HMI tags "Default tag table"
   "Clock_0.5Hz" : Bool = PLC "Clock_0.5Hz", 1 s
   "messageView" : Bool, internal
   "buttonView" : Bool, internal
   "RPA10B_datablock_PA10B_fatal_error_state_lock" : Int, 1 s
   "RPA10B_datablock_PA10B_error_state_lock" : Int, 1 s
   "RPA10B_datablock_PA10B_big_fail_state_lock" : Int, 1 s
   "RPA10B_datablock_PA10B_fail_state_lock" : Int, 1 s
   "RPA10B_datablock_RPA10B_station_work_cyclus_state" : UInt, 1 s
   "RPA10R_LCDSwitchAutomat_Manual" : Bool = PLC "RPA10B_LCD_switch_manual_automat", 1 s
   "RPA10B_datablock_RPA10B_station_start" : Bool, 1 s
   "show_input_page" : Int, internal
   "PLC_datablock_stations_configuration" : Byte, 1 s
   "RPA10B_datablock_RPA10B_instruction_list_index" : Byte, 1 s
   "RPA20B_open_drawer" : Bool = PLC "RPA20B_open_drawer", 1 s
   "RPA10B_LCD_switch_manual_automat" : Bool = PLC "RPA10B_LCD_switch_manual_automat", 1 s
   "RPA10B_datablock_RPA10B_scanned_data" : String[254], 1 s
   "RPA10B_light" : Bool = PLC "RPA10B_light", 1 s
   "RPA10B_LCD_beacon_green" : Bool = PLC "RPA10B_LCD_beacon_green", 1 s
   "RPA10B_LCD_beacon_orange" : Bool = PLC "RPA10B_LCD_beacon_orange", 1 s
   "RPA10B_LCD_beacon_red" : Bool = PLC "RPA10B_LCD_beacon_red", 1 s
   "RPA10B_LCD_beacon_siren" : Bool = PLC "RPA10B_LCD_beacon_siren", 1 s
   "RPA10B_LCD_button_start" : Bool = PLC "RPA10B_LCD_button_start", 1 s
   "RPA10B_LCD_LED_blue_confirm_button" : Bool = PLC "RPA10B_LCD_LED_blue_confirm_button", 1 s
   "RPA10B_LCD_LED_green_start_button" : Bool = PLC "RPA10B_LCD_LED_green_start_button", 1 s
   "RPA10B_code_position_1" : Bool = PLC "RPA10B_code_position_1", 1 s
   "RPA10B_code_position_2" : Bool = PLC "RPA10B_code_position_2", 1 s
   "RPA10B_home_position_horizontal_carriage_sensor" : Bool = PLC "RPA10B_home_position_horizontal_carriage_sensor", 1 s
   "RPA10B_end_position_horizontal_carriage_sensor" : Bool = PLC "RPA10B_end_position_horizontal_carriage_sensor", 1 s
   "RPA10B_home_position_idler_carriage_sensor" : Bool = PLC "RPA10B_home_position_idler_carriage_sensor", 1 s
   "RPA10B_end_position_idler_carriage_sensor" : Bool = PLC "RPA10B_end_position_idler_carriage_sensor", 1 s
   "RPA10B_idler_presence_sensor" : Bool = PLC "RPA10B_idler_presence_sensor", 1 s
   "show_output_page" : Int, internal
   "input_output" : Bool, internal
   "RPA10B_vacuum_sensor" : Bool = PLC "RPA10B_vacuum_sensor", 1 s
   "RPA10B_lock_sensor" : Bool = PLC "RPA10B_lock_sensor", 1 s
   "RPA10B_unlock_sensor" : Bool = PLC "RPA10B_unlock_sensor", 1 s
   "RPA10B_blend_1_vacuum_fix_sensor" : Bool = PLC "RPA10B_blend_1_vacuum_fix_sensor", 1 s
   "RPA10B_blend_2_vacuum_fix_sensor" : Bool = PLC "RPA10B_blend_2_vacuum_fix_sensor", 1 s
   "RPA10B_LCD_button_confirm" : Bool = PLC "RPA10B_LCD_button_confirm", 1 s
   "RPA10B_primerbox_pad_sensor_left" : Bool = PLC "RPA10B_primerbox_pad_sensor_left", 1 s
   "RPA10B_primerbox_pad_sensor_right" : Bool = PLC "RPA10B_primerbox_pad_sensor_right", 1 s
   "RPA10B_primerbox_felt_sensor" : Bool = PLC "RPA10B_primerbox_felt_sensor", 1 s
   "RPA10B_primerbox_felt_presence_sensor" : Bool = PLC "RPA10B_primerbox_felt_presence_sensor", 1 s
   "RPA10B_primerbox_button_PAD_IS_CHANGED" : Bool = PLC "RPA10B_primerbox_button_PAD_IS_CHANGED", 1 s
   "RPA10B_primerbox_bottle_2" : Bool = PLC "RPA10B_primerbox_bottle_2", 1 s
   "RPA10B_primerbox_bottle_1" : Bool = PLC "RPA10B_primerbox_bottle_1", 1 s
   "RPA10B_EJ_1_vacuum_sensor" : Bool = PLC "RPA10B_EJ_1_vacuum_sensor", 1 s
   "RPA10B_EJ_2_vacuum_sensor" : Bool = PLC "RPA10B_EJ_2_vacuum_sensor", 1 s
   "RPA10B_universal_button_1" : Bool = PLC "RPA10B_universal_button_1", 1 s
   "RPA10B_universal_button_2" : Bool = PLC "RPA10B_universal_button_2", 1 s
   "RPA20B_belt_position_sensor" : Bool = PLC "RPA20B_belt_position_sensor", 1 s
   "RPA20B_blend_presence_sensor_1" : Bool = PLC "RPA20B_blend_presence_sensor_1", 1 s
   "RPA20B_blend_presence_sensor_2" : Bool = PLC "RPA20B_blend_presence_sensor_2", 1 s
   "RPA20B_drawer_position_sensor" : Bool = PLC "RPA20B_drawer_position_sensor", 1 s
   "RPA20B_drawer_lock_sensor" : Bool = PLC "RPA20B_drawer_lock_sensor", 1 s
   "RPA20B_drawer_unlock_sensor" : Bool = PLC "RPA20B_drawer_unlock_sensor", 1 s
   "RPA20B_ES_feedback" : Bool = PLC "RPA20B_ES_feedback", 1 s
   "RPA20B_lock_door_feedback" : Bool = PLC "RPA20B_lock_door_feedback", 1 s
   "RPA20B_manual_UP" : Bool = PLC "RPA20B_manual_UP", 1 s
   "RPA20B_manual_DOWN" : Bool = PLC "RPA20B_manual_DOWN", 1 s
   "RPA20B_manual_move" : Bool = PLC "RPA20B_manual_move", 1 s
   "RPA20B_unlock_button" : Bool = PLC "RPA20B_unlock_button", 1 s
   "RPA20B_button_back_1" : Bool = PLC "RPA20B_button_back_1", 1 s
   "RPA20B_button_back_2" : Bool = PLC "RPA20B_button_back_2", 1 s
   "RPA10B_primerbox_beacon_green" : Bool = PLC "RPA10B_primerbox_beacon_green", 1 s
   "RPA10B_primerbox_beacon_orange" : Bool = PLC "RPA10B_primerbox_beacon_orange", 1 s
   "RPA10B_primerbox_beacon_red" : Bool = PLC "RPA10B_primerbox_beacon_red", 1 s
   "RPA10B_primerbox_beacon_siren" : Bool = PLC "RPA10B_primerbox_beacon_siren", 1 s
   "RPA10B_primerbox_LED_green_ready" : Bool = PLC "RPA10B_primerbox_LED_green_ready", 1 s
   "RPA10B_primerbox_LED_green_felt" : Bool = PLC "RPA10B_primerbox_LED_green_felt", 1 s
   "RPA10B_primerbox_LED_green_bottle_1" : Bool = PLC "RPA10B_primerbox_LED_green_bottle_1", 1 s
   "RPA10B_primerbox_LED_green_bottle_2" : Bool = PLC "RPA10B_primerbox_LED_green_bottle_2", 1 s
   "RPA10B_primerbox_LED_red_NOT_READY" : Bool = PLC "RPA10B_primerbox_LED_red_NOT_READY", 1 s
   "RPA10B_primerbox_LED_orange_change_pad" : Bool = PLC "RPA10B_primerbox_LED_orange_change_pad", 1 s
   "RPA10B_vavle_aretation_unlock" : Bool = PLC "RPA10B_vavle_aretation_unlock", 1 s
   "RPA10B_vavle_aretation_lock" : Bool = PLC "RPA10B_vavle_aretation_lock", 1 s
   "RPA10B_vavle_seal_idler_unlock" : Bool = PLC "RPA10B_vavle_seal_idler_unlock", 1 s
   "RPA10B_vavle_seal_idler_lock" : Bool = PLC "RPA10B_vavle_seal_idler_lock", 1 s
   "RPA10B_EJ_1_vacuum_control" : Bool = PLC "RPA10B_EJ_1_vacuum_control", 1 s
   "RPA10B_EJ_2_vacuum_control" : Bool = PLC "RPA10B_EJ_2_vacuum_control", 1 s
   "RPA10B_EJ_1_eject" : Bool = PLC "RPA10B_EJ_1_eject", 1 s
   "RPA10B_EJ_2_eject" : Bool = PLC "RPA10B_EJ_2_eject", 1 s
   "RPA10B_vacuum_cleaner_switch" : Bool = PLC "RPA10B_vacuum_cleaner_switch", 1 s
   "RPA20B_open_door_LED_green" : Bool = PLC "RPA20B_open_door_LED_green", 1 s
   "RPA20B_button_back_LED_1" : Bool = PLC "RPA20B_button_back_LED_1", 1 s
   "RPA20B_button_back_LED_2" : Bool = PLC "RPA20B_button_back_LED_2", 1 s
   "RPA20B_valve_open_drawer" : Bool = PLC "RPA20B_valve_open_drawer", 1 s
   "RPA20B_valve_close_drawer" : Bool = PLC "RPA20B_valve_close_drawer", 1 s
   "RPA20B_motor_down" : Bool = PLC "RPA20B_motor_down", 1 s
   "RPA20_motor_up" : Bool = PLC "RPA20_motor_up", 1 s
   "manual_page_switch" : Int, internal
   "RPA10B_datablock_RPA10B_show_pad_left" : Bool, 1 s
   "RPA10B_datablock_RPA10B_show_pad_right" : Bool, 1 s
   "RPA10B_datablock_RPA10_B_show_home" : Bool, 1 s
   "RPA10B_datablock_pa10B_bottle_cyclus_replace" : UInt, 1 s
   "RPA10B_datablock_pa10B_bottle_timing" : Time, 1 s

text list "PA10B_instructionList": 0 ''; 1 ''; 2 ''; 4 ''; 6 ''; 7 ''; 8 ''; 3 ''; 5 ''; 9 ''; 11 ''; 12 ''; 13 ''; 14 ''; 15 ''; 16 ''; 17 ''; 18 ''; 19 ''; 20 ''; 21 ''; 22 ''; 23 ''; 24 ''; 25 ''; 26 ''; 27 ''; 28 ''; 29 ''; 30 ''; 31 ''; 70 ''

text list "PA10B_fatal_error_list": 150 ''; 1100 ''

text list "pa10B_fail_list": 150 ''; 303 ''; 304 ''; 203 ''; 204 ''; 205 ''; 180 ''

text list "PA10B_error_list": 1000 ''; 400 ''; 401 ''; 402 ''; 403 ''

text list "PA10B_big_fail_list": 305 ''; 205 ''; 169 ''

text list "PA10B_station_variant_choose": 0 ''; 1 ''; 2 ''; 3 ''

screen "Home" 800x480
   TextField "Text field_3" at 325,5 size 300x40
   TextField "Text field_2" at 2,85 size 70x40
   TextField "Text field_5" at 335,130 size 130x25
   TextField "Text field_6" at 20,171 size 330x22
   TextField "Text field_7" at 20,201 size 330x22
   TextField "Text field_8" at 20,231 size 330x22
   TextField "Text field_9" at 20,261 size 330x22
   TextField "Text field_10" at 20,291 size 330x22
   TextField "Text field_11" at 20,321 size 330x22
   TextField "Text field_12" at 20,351 size 330x22
   TextField "Text field_13" at 20,381 size 330x22
   Button "Button_1" at 640,420 size 80x60
   Button "HmiScreenItemData_1" at 0,420 size 80x60
   Button "HmiScreenItemData_2" at 400,420 size 80x60
   Button "Button_2" at 560,420 size 80x60
   Button "Button_6" at 720,420 size 80x60
   DateTimeField "Date/time field_1" at 650,27 size 150x25
   DateTimeField "Date/time field_2" at 650,0 size 150x28
   TextField "Text field_1" at 0,0 size 300x50
   Button "HmiScreenItemData_3" at 240,420 size 80x60
   Button "HmiScreenItemData_4" at 320,420 size 80x60
   Button "Button_3" at 480,420 size 80x60
   Button "HmiScreenItemData_5" at 80,420 size 80x60
   Button "HmiScreenItemData_6" at 160,420 size 80x60
   IOField "I/O field_1" at 73,85 size 70x40
   Button "Button_11" at 0,420 size 80x60
   Button "Button_12" at 80,420 size 80x60
   Button "Button_13" at 160,420 size 80x60
   Button "Button_14" at 240,420 size 80x60
   Button "Button_15" at 320,420 size 80x60
   Button "Button_16" at 400,420 size 80x60
   Button "Button_17" at 480,420 size 80x60
   Button "Button_18" at 560,420 size 80x60
   Button "Button_19" at 640,420 size 80x60
   Button "Button_20" at 720,420 size 80x60
   TextField "Text field_22" at 64,67 size 129x22
   AlarmView "Alarm view_1" at 60,90 size 680x320
   Button "Button_9" at 715,65 size 25x25
   TextField "Text field_37" at 360,54 size 120x25

screen "I0-State" 800x480
   TextField "Text field_3" at 325,5 size 300x40
   Button "Button_1" at 640,420 size 80x60
   Button "Button_4" at 160,420 size 80x60
   Button "HmiScreenItemData_3" at 400,420 size 80x60
   Button "Button_2" at 560,420 size 80x60
   Button "Button_6" at 720,420 size 80x60
   Button "HmiScreenItemData_2" at 240,420 size 80x60
   Button "HmiScreenItemData_4" at 320,420 size 80x60
   TextField "Text field_1" at 0,0 size 300x50
   DateTimeField "Date/time field_2" at 650,0 size 150x28
   DateTimeField "Date/time field_1" at 650,27 size 150x25
   Button "HmiScreenItemData_1" at 0,420 size 80x60
   Button "Button_3" at 480,420 size 80x60
   Button "Button_5" at 80,420 size 80x60
   Button "input_back" at 20,52 size 90x25
   Button "input_next" at 690,52 size 90x25
   Button "output_back" at 20,52 size 90x25
   Button "output_next" at 690,52 size 90x25
   TextField "Text field_2" at 20,85 size 330x22
   TextField "Text field_4" at 20,114 size 330x22
   TextField "Text field_5" at 20,144 size 330x22
   TextField "Text field_6" at 20,174 size 330x22
   TextField "Text field_13" at 20,204 size 330x22
   TextField "Text field_14" at 20,232 size 330x22
   TextField "Text field_15" at 20,260 size 330x22
   TextField "Text field_16" at 20,288 size 330x22
   TextField "Text field_17" at 20,316 size 330x22
   TextField "Text field_18" at 20,344 size 330x22
   TextField "Text field_19" at 19,374 size 330x22
   TextField "Text field_20" at 387,86 size 330x22
   TextField "Text field_21" at 387,115 size 330x22
   TextField "Text field_22" at 387,144 size 330x22
   TextField "Text field_23" at 387,173 size 330x22
   TextField "Text field_24" at 387,202 size 330x22
   TextField "Text field_26" at 387,231 size 330x22
   TextField "Text field_27" at 387,260 size 330x22
   TextField "Text field_28" at 387,289 size 330x22
   TextField "Text field_29" at 387,318 size 330x22
   TextField "Text field_30" at 387,347 size 330x22
   TextField "Text field_31" at 387,376 size 330x22
   Button "Button_11" at 0,420 size 80x60
   Button "Button_12" at 80,420 size 80x60
   Button "Button_13" at 160,420 size 80x60
   Button "Button_14" at 240,420 size 80x60
   Button "Button_15" at 320,420 size 80x60
   Button "Button_16" at 400,420 size 80x60
   Button "Button_17" at 480,420 size 80x60
   Button "Button_18" at 560,420 size 80x60
   Button "Button_19" at 640,420 size 80x60
   Button "Button_20" at 720,420 size 80x60
   TextField "Text field_25" at 64,67 size 129x22
   AlarmView "Alarm view_1" at 60,90 size 680x320
   Button "Button_9" at 715,65 size 25x25
   TextField "Text field_7" at 20,85 size 330x22
   TextField "Text field_8" at 19,115 size 330x22
   TextField "Text field_9" at 19,145 size 330x22
   TextField "Text field_10" at 19,175 size 330x22
   TextField "Text field_11" at 20,205 size 330x22
   TextField "Text field_12" at 20,235 size 330x22
   TextField "Text field_50" at 20,263 size 330x22
   TextField "Text field_51" at 20,291 size 330x22
   TextField "Text field_52" at 20,319 size 330x22
   TextField "Text field_53" at 20,347 size 330x22
   TextField "Text field_54" at 20,375 size 330x22
   TextField "Text field_55" at 387,86 size 330x22
   TextField "Text field_56" at 386,116 size 330x22
   TextField "Text field_57" at 386,146 size 330x22
   TextField "Text field_58" at 386,176 size 330x22
   TextField "Text field_59" at 387,206 size 330x22
   TextField "Text field_60" at 387,236 size 330x22
   TextField "Text field_61" at 387,264 size 330x22
   TextField "Text field_62" at 387,292 size 330x22
   TextField "Text field_63" at 387,320 size 330x22
   TextField "Text field_64" at 387,348 size 330x22
   TextField "Text field_65" at 387,376 size 330x22
   TextField "Text field_32" at 20,85 size 330x22
   TextField "Text field_33" at 20,114 size 330x22
   TextField "Text field_34" at 20,144 size 330x22
   TextField "Text field_35" at 20,174 size 330x22
   TextField "Text field_36" at 20,204 size 330x22
   TextField "Text field_37" at 20,232 size 330x22
   TextField "Text field_38" at 20,260 size 330x22
   TextField "Text field_39" at 20,288 size 330x22
   TextField "Text field_40" at 20,316 size 330x22
   TextField "Text field_41" at 20,344 size 330x22
   TextField "Text field_42" at 19,374 size 330x22
   TextField "Text field_43" at 387,86 size 330x22
   TextField "Text field_44" at 387,115 size 330x22
   TextField "Text field_45" at 387,144 size 330x22
   TextField "Text field_46" at 387,173 size 330x22
   TextField "Text field_47" at 387,202 size 330x22
   TextField "Text field_48" at 387,231 size 330x22
   TextField "Text field_49" at 387,260 size 330x22
   TextField "Text field_66" at 20,85 size 330x22
   TextField "Text field_67" at 19,115 size 330x22
   TextField "Text field_68" at 19,145 size 330x22
   TextField "Text field_69" at 19,175 size 330x22
   TextField "Text field_70" at 20,205 size 330x22
   TextField "Text field_71" at 20,235 size 330x22
   TextField "Text field_72" at 20,263 size 330x22
   TextField "Text field_73" at 20,291 size 330x22
   TextField "Text field_74" at 20,319 size 330x22
   TextField "Text field_75" at 20,347 size 330x22
   TextField "Text field_76" at 20,375 size 330x22
   TextField "Text field_77" at 360,54 size 120x25

screen "Main_page" 800x480
   Button "HmiScreenItemData_1" at 80,420 size 80x60
   TextField "Text field_2" at 0,85 size 800x25
   TextField "Text field_3" at 325,5 size 300x40
   Button "Button_4" at 480,420 size 80x60
   Button "Button_5" at 640,420 size 80x60
   Button "Button_1" at 0,420 size 80x60
   Button "HmiScreenItemData_2" at 160,420 size 80x60
   Button "Button_2" at 400,420 size 80x60
   Button "Button_3" at 560,420 size 80x60
   Button "Button_6" at 720,420 size 80x60
   Button "HmiScreenItemData_3" at 240,420 size 80x60
   Button "HmiScreenItemData_4" at 320,420 size 80x60
   TextField "Text field_1" at 0,0 size 300x50
   DateTimeField "Date/time field_2" at 650,0 size 150x28
   DateTimeField "Date/time field_1" at 650,27 size 150x25
   SymbolicIOField "Symbolic I/O field_1" at 10,110 size 780x90
   Button "HmiScreenItemData_5" at 80,420 size 80x60
   GraphicView "Graphic view_1" at 320,228 size 180x180
   Button "Button_11" at 0,420 size 80x60
   Button "Button_12" at 80,420 size 80x60
   Button "Button_13" at 160,420 size 80x60
   Button "Button_14" at 240,420 size 80x60
   Button "Button_15" at 320,420 size 80x60
   Button "Button_16" at 400,420 size 80x60
   Button "Button_17" at 480,420 size 80x60
   Button "Button_18" at 560,420 size 80x60
   Button "Button_19" at 640,420 size 80x60
   Button "Button_20" at 720,420 size 80x60
   TextField "Text field_5" at 64,67 size 129x22
   AlarmView "Alarm view_1" at 60,90 size 680x320
   Button "Button_9" at 715,65 size 25x25
   SymbolicIOField "Symbolic I/O field_2" at 0,170 size 800x110
   SymbolicIOField "Symbolic I/O field_3" at 0,170 size 800x110
   SymbolicIOField "Symbolic I/O field_4" at 0,170 size 800x110
   SymbolicIOField "Symbolic I/O field_5" at 0,170 size 800x110
   TextField "Text field_37" at 360,54 size 120x25
   GraphicView "Graphic view_2" at 260,225 size 345x187
   GraphicView "Graphic view_3" at 195,225 size 345x187
   TextField "Text field_4" at 306,290 size 237x43

screen "Manual" 800x480
   Button "Button_4" at 21,85 size 50x50
   Button "Button_12" at 730,85 size 50x50
   Button "Button_1" at 640,420 size 80x60
   Button "HmiScreenItemData_1" at 0,420 size 80x60
   Button "Button_2" at 560,420 size 80x60
   Button "Button_6" at 720,420 size 80x60
   Button "Button_34" at 400,420 size 80x60
   Button "HmiScreenItemData_3" at 240,420 size 80x60
   Button "HmiScreenItemData_4" at 320,420 size 80x60
   TextField "Text field_1" at 0,0 size 300x50
   DateTimeField "Date/time field_2" at 650,0 size 150x28
   DateTimeField "Date/time field_1" at 650,27 size 150x25
   Button "Button_5" at 160,420 size 80x60
   Button "Button_3" at 480,420 size 80x60
   Button "Button_7" at 80,420 size 80x60
   Button "Button_8" at 730,85 size 50x50
   Button "Button_9" at 21,85 size 50x50
   Button "Button_23" at 0,420 size 80x60
   Button "Button_24" at 80,420 size 80x60
   Button "Button_25" at 160,420 size 80x60
   Button "Button_26" at 240,420 size 80x60
   Button "Button_27" at 320,420 size 80x60
   Button "Button_28" at 400,420 size 80x60
   Button "Button_29" at 480,420 size 80x60
   Button "Button_30" at 560,420 size 80x60
   Button "Button_31" at 640,420 size 80x60
   Button "Button_32" at 720,420 size 80x60
   TextField "Text field_8" at 64,67 size 129x22
   AlarmView "Alarm view_1" at 60,90 size 680x320
   Button "Button_33" at 715,65 size 25x25
   Switch "Switch_8" at 300,149 size 64x32
   Switch "Switch_9" at 300,185 size 64x32
   Switch "Switch_10" at 300,221 size 64x32
   Switch "Switch_11" at 300,257 size 64x32
   Switch "Switch_12" at 300,293 size 64x32
   Switch "Switch_13" at 301,328 size 64x32
   TextField "Text field_15" at 76,149 size 200x32
   TextField "Text field_16" at 76,181 size 200x32
   TextField "Text field_17" at 75,221 size 200x32
   TextField "Text field_18" at 37,289 size 239x32
   TextField "Text field_19" at 26,257 size 250x32
   TextField "Text field_20" at 29,328 size 247x32
   Switch "Switch_1" at 634,148 size 64x32
   TextField "Text field_2" at 410,148 size 200x32
   Switch "Switch_2" at 301,363 size 64x32
   TextField "Text field_4" at 29,363 size 247x32
   Switch "Switch_3" at 634,184 size 64x32
   TextField "Text field_5" at 379,184 size 231x32
   Switch "Switch_4" at 635,220 size 64x32
   TextField "Text field_6" at 394,220 size 217x32
   Switch "Switch_5" at 636,256 size 64x32
   TextField "Text field_7" at 377,256 size 235x32
   Switch "Switch_6" at 637,292 size 64x32
   TextField "Text field_9" at 377,292 size 236x32
   Switch "Switch_7" at 638,328 size 64x32
   TextField "Text field_10" at 376,328 size 238x32
   Switch "Switch_14" at 639,364 size 64x32
   TextField "Text field_11" at 322,364 size 293x32
   Switch "Switch_15" at 300,149 size 64x32
   Switch "Switch_16" at 300,185 size 64x32
   Switch "Switch_17" at 300,221 size 64x32
   Switch "Switch_18" at 300,257 size 64x32
   Switch "Switch_19" at 300,293 size 64x32
   Switch "Switch_20" at 301,328 size 64x32
   TextField "Text field_12" at 55,149 size 221x32
   TextField "Text field_13" at 8,181 size 268x32
   TextField "Text field_14" at 44,221 size 231x32
   TextField "Text field_21" at 37,289 size 239x32
   TextField "Text field_22" at 26,257 size 250x32
   TextField "Text field_23" at 29,328 size 247x32
   Switch "Switch_21" at 634,148 size 64x32
   TextField "Text field_24" at 388,148 size 222x32
   Switch "Switch_22" at 301,363 size 64x32
   TextField "Text field_25" at 29,363 size 247x32
   Switch "Switch_23" at 634,184 size 64x32
   TextField "Text field_26" at 379,184 size 231x32
   Switch "Switch_24" at 635,220 size 64x32
   TextField "Text field_27" at 394,220 size 217x32
   Switch "Switch_25" at 636,256 size 64x32
   TextField "Text field_28" at 377,256 size 235x32
   Switch "Switch_26" at 637,292 size 64x32
   TextField "Text field_29" at 377,292 size 236x32
   Switch "Switch_27" at 638,328 size 64x32
   TextField "Text field_30" at 376,328 size 238x32
   Switch "Switch_28" at 639,364 size 64x32
   TextField "Text field_31" at 382,364 size 233x32
   Switch "Switch_29" at 300,149 size 64x32
   Switch "Switch_30" at 300,185 size 64x32
   Switch "Switch_31" at 300,221 size 64x32
   Switch "Switch_32" at 300,257 size 64x32
   Switch "Switch_33" at 300,293 size 64x32
   TextField "Text field_32" at 55,149 size 221x32
   TextField "Text field_33" at 8,181 size 268x32
   TextField "Text field_34" at 22,221 size 253x32
   TextField "Text field_35" at 37,289 size 239x32
   TextField "Text field_36" at 26,257 size 250x32
   TextField "Text field_37" at 360,54 size 120x25

screen "Scanner" 800x480
   IOField "I/O field_1" at 10,118 size 780x32
   TextField "Text field_2" at 10,86 size 141x22
   Button "Button_1" at 640,420 size 80x60
   Button "HmiScreenItemData_3" at 400,420 size 80x60
   Button "Button_2" at 560,420 size 80x60
   Button "Button_6" at 720,420 size 80x60
   DateTimeField "Date/time field_2" at 650,0 size 150x28
   TextField "Text field_1" at 0,0 size 300x50
   DateTimeField "Date/time field_1" at 650,27 size 150x25
   Button "HmiScreenItemData_2" at 240,420 size 80x60
   Button "HmiScreenItemData_4" at 320,420 size 80x60
   Button "HmiScreenItemData_1" at 0,420 size 80x60
   Button "HmiScreenItemData_5" at 480,420 size 80x60
   Button "HmiScreenItemData_6" at 160,420 size 80x60
   Button "HmiScreenItemData_7" at 80,420 size 80x60
   Button "Button_3" at 10,170 size 96x32
   Button "Button_11" at 0,420 size 80x60
   Button "Button_12" at 80,420 size 80x60
   Button "Button_13" at 160,420 size 80x60
   Button "Button_14" at 240,420 size 80x60
   Button "Button_15" at 320,420 size 80x60
   Button "Button_16" at 400,420 size 80x60
   Button "Button_17" at 480,420 size 80x60
   Button "Button_18" at 560,420 size 80x60
   Button "Button_19" at 640,420 size 80x60
   Button "Button_20" at 720,420 size 80x60
   TextField "Text field_5" at 64,67 size 129x22
   Button "Button_9" at 715,65 size 25x25
   AlarmView "Alarm view_1" at 60,90 size 680x320
   TextField "Text field_37" at 360,54 size 120x25

screen "System" 800x480
   TextField "Text field_3" at 325,5 size 300x40
   TextField "Text field_2" at 300,85 size 200x27
   Button "Button_4" at 10,290 size 170x60
   Button "Button_5" at 10,355 size 170x60
   Button "Button_7" at 213,290 size 170x60
   Button "Button_8" at 416,290 size 170x60
   Button "Button_9" at 620,290 size 170x60
   Button "Button_11" at 213,355 size 170x60
   Button "Button_12" at 416,355 size 170x60
   Button "Button_13" at 620,355 size 170x60
   AlarmView "Alarm view_1" at 10,113 size 780x172
   Button "HmiScreenItemData_1" at 0,420 size 80x60
   Button "Button_3" at 160,420 size 80x60
   Button "Button_14" at 240,420 size 80x60
   Button "Button_15" at 320,420 size 80x60
   Button "Button_16" at 400,420 size 80x60
   Button "Button_17" at 480,420 size 80x60
   Button "Button_2" at 560,420 size 80x60
   Button "Button_1" at 640,420 size 80x60
   Button "Button_6" at 720,420 size 80x60
   TextField "Text field_1" at 0,0 size 300x50
   DateTimeField "Date/time field_2" at 650,0 size 150x28
   DateTimeField "Date/time field_1" at 650,27 size 150x25
   Button "Button_10" at 80,420 size 80x60
   TextField "Text field_37" at 360,54 size 120x25

screen "chemical_setup" 800x480
   Button "HmiScreenItemData_3" at 400,420 size 80x60
   Button "Button_2" at 560,420 size 80x60
   Button "Button_6" at 720,420 size 80x60
   DateTimeField "Date/time field_2" at 650,0 size 150x28
   TextField "Text field_1" at 0,0 size 300x50
   DateTimeField "Date/time field_1" at 650,27 size 150x25
   Button "HmiScreenItemData_2" at 240,420 size 80x60
   Button "HmiScreenItemData_4" at 320,420 size 80x60
   Button "HmiScreenItemData_1" at 0,420 size 80x60
   Button "HmiScreenItemData_5" at 480,420 size 80x60
   Button "HmiScreenItemData_6" at 160,420 size 80x60
   Button "HmiScreenItemData_7" at 80,420 size 80x60
   IOField "I/O field_1" at 87,130 size 341x44
   IOField "I/O field_2" at 87,237 size 338x44
   TextField "Text field_2" at 85,100 size 137x25
   TextField "Text field_3" at 87,206 size 111x25
   TextField "Text field_4" at 435,245 size 93x20
   Button "Button_1" at 640,420 size 80x60
   Button "Button_11" at 0,420 size 80x60
   Button "Button_12" at 80,420 size 80x60
   Button "Button_13" at 160,420 size 80x60
   Button "Button_14" at 240,420 size 80x60
   Button "Button_15" at 320,420 size 80x60
   Button "Button_16" at 400,420 size 80x60
   Button "Button_17" at 480,420 size 80x60
   Button "Button_18" at 560,420 size 80x60
   Button "Button_19" at 640,420 size 80x60
   Button "Button_20" at 720,420 size 80x60
   TextField "Text field_5" at 64,67 size 129x22
   Button "Button_9" at 715,65 size 25x25
   AlarmView "Alarm view_1" at 60,90 size 680x320
   TextField "Text field_37" at 360,54 size 120x25

screen "User_management" 800x480
   TextField "Text field_3" at 325,5 size 300x40
   Button "HmiScreenItemData_1" at 0,420 size 80x60
   Button "Button_3" at 160,420 size 80x60
   Button "Button_14" at 240,420 size 80x60
   Button "Button_15" at 320,420 size 80x60
   Button "Button_16" at 400,420 size 80x60
   Button "Button_17" at 480,420 size 80x60
   Button "Button_2" at 560,420 size 80x60
   Button "Button_1" at 640,420 size 80x60
   TextField "Text field_1" at 0,0 size 300x50
   DateTimeField "Date/time field_2" at 650,0 size 150x28
   DateTimeField "Date/time field_1" at 650,27 size 150x25
   Button "Button_10" at 80,420 size 80x60
   UserView "User view_1" at 20,92 size 758x304
   Button "Button_4" at 720,420 size 80x60
   TextField "Text field_37" at 360,54 size 120x25
*)

(* ===== HMI "HMI_RT_7" =====
connection "HMI_Connection_6": ETHERNET, SMART_S7_1500_OMS

HMI tags "Default tag table"
   "Clock_0.5Hz" : Bool = PLC "Clock_0.5Hz", 1 s
   "FS_datablock_fs_alarm" : Bool, 1 s
   "fs_datablock_fs_chemical_type" : Byte, 100 ms
   "FS_datablock_fs_error_identifier" : Int, 1 s
   "fs_datablock_fs_expire_time_Activator_DW646" : DInt, 1 s
   "fs_datablock_fs_expire_time_Activator_SIKA_110" : DInt, 1 s
   "fs_datablock_fs_expire_time_Primer_DV954V1" : DInt, 1 s
   "fs_datablock_fs_expire_time_Primer_SIKA_207" : DInt, 1 s
   "fs_datablock_fs_expire_time_Remover_SIKA_208" : DInt, 1 s
   "fs_datablock_fs_filling_e" : Bool, 1 s
   "fs_datablock_fs_funel_control{1}" : Bool, 1 s
   "fs_datablock_fs_funel_control{2}" : Bool, 1 s
   "fs_datablock_fs_funel_control{3}" : Bool, 1 s
   "fs_datablock_fs_funel_control{4}" : Bool, 1 s
   "fs_datablock_fs_funel_control{5}" : Bool, 1 s
   "FS_datablock_fs_hmi_instruction_index" : Byte, 100 ms
   "fs_datablock_fs_input_expire_date" : USInt, 1 s
   "fs_datablock_fs_input_expire_year" : UInt, 1 s
   "fs_datablock_fs_mixer_expiration_sec{0}" : Int, 1 s
   "fs_datablock_fs_mixer_expiration_sec{1}" : Int, 1 s
   "fs_datablock_fs_mixer_expiration_sec{2}" : Int, 1 s
   "fs_datablock_fs_mixer_expiration_sec{3}" : Int, 1 s
   "fs_datablock_fs_mixer_expiration_sec{4}" : Int, 1 s
   "fs_datablock_fs_primer_DV954V1_shake_time" : Time, 1 s
   "fs_datablock_fs_primer_DV954V1_time_after_shaking" : Time, 1 s
   "fs_datablock_fs_primer_SIKA_207_shake_time" : Time, 1 s
   "fs_datablock_fs_primer_SIKA_207_time_after_shaking" : Time, 1 s
   "fs_datablock_fs_print_sp_bottle_e" : Bool, 1 s
   "fs_datablock_fs_reset_e" : Bool, 1 s
   "FS_datablock_fs_scaned_data" : String[254], 1 s
   "fs_datablock_fs_shaker_batch_code_str{0}" : String[254], 1 s
   "fs_datablock_fs_shaker_batch_code_str{1}" : String[254], 1 s
   "fs_datablock_fs_shaker_batch_code_str{2}" : String[254], 1 s
   "fs_datablock_fs_shaker_batch_code_str{3}" : String[254], 1 s
   "fs_datablock_fs_shaker_batch_code_str{4}" : String[254], 1 s
   "fs_datablock_fs_shaker_chemical_type_str{0}" : String[254], 1 s
   "fs_datablock_fs_shaker_chemical_type_str{1}" : String[254], 1 s
   "fs_datablock_fs_shaker_chemical_type_str{2}" : String[254], 1 s
   "fs_datablock_fs_shaker_chemical_type_str{3}" : String[254], 1 s
   "fs_datablock_fs_shaker_chemical_type_str{4}" : String[254], 1 s
   "fs_datablock_fs_shaker_expiration_str{0}" : String[254], 1 s
   "fs_datablock_fs_shaker_expiration_str{1}" : String[254], 1 s
   "fs_datablock_fs_shaker_expiration_str{2}" : String[254], 1 s
   "fs_datablock_fs_shaker_expiration_str{3}" : String[254], 1 s
   "fs_datablock_fs_shaker_expiration_str{4}" : String[254], 1 s
   "FS_datablock_fs_show_button" : Bool, 100 ms
   "fs_datablock_fs_show_fill_button{1}" : Bool, 1 s
   "fs_datablock_fs_show_fill_button{2}" : Bool, 1 s
   "fs_datablock_fs_show_fill_button{3}" : Bool, 1 s
   "fs_datablock_fs_show_fill_button{4}" : Bool, 1 s
   "fs_datablock_fs_show_fill_button{5}" : Bool, 1 s
   "FS_datablock_fs_statin_activity_state" : Bool, 1 s
   "fs_fill_bottle_fce_DB_chemical_type" : Byte, 1 s
   "FS_LCD_button_confirm" : Bool = PLC "ib_FS_LCD_button_confirm", 1 s
   "FS_LCD_button_start" : Bool = PLC "ib_FS_LCD_button_start", 1 s
   "FS_LCD_confirm_button_LED_blue" : Bool = PLC "ob_FS_LCD_confirm_button_LED_blue", 5 s
   "FS_LCD_start_button_LED_green" : Bool = PLC "ob_FS_LCD_start_button_LED_green", 5 s
   "FS_move_UP_funel_1" : Bool = PLC "ob_FS_move_UP_funel_1"
   "FS_move_UP_funel_2" : Bool = PLC "ob_FS_move_UP_funel_2"
   "FS_move_UP_funel_3" : Bool = PLC "ob_FS_move_UP_funel_3"
   "FS_move_UP_funel_4" : Bool = PLC "ob_FS_move_UP_funel_4"
   "FS_move_UP_funel_5" : Bool = PLC "ob_FS_move_UP_funel_5"
   "fs_print_lable_suplier_bottle_DB_batch_code" : String[254], 1 s
   "fs_print_lable_suplier_bottle_DB_chemical_code" : String[254], 1 s
   "FS_sensor_bottle_1" : Bool = PLC "ib_FS_sensor_bottle_1", 5 s
   "FS_sensor_bottle_2" : Bool = PLC "ib_FS_sensor_bottle_2", 5 s
   "FS_sensor_bottle_3" : Bool = PLC "ib_FS_sensor_bottle_3", 5 s
   "FS_sensor_bottle_4" : Bool = PLC "ib_FS_sensor_bottle_4", 5 s
   "FS_sensor_bottle_5" : Bool = PLC "ib_FS_sensor_bottle_5", 5 s
   "ib_FS_LCD_switch_automat_manual" : Bool = PLC "ib_FS_LCD_switch_automat_manual", 1 s
   "ib_FS_mixer_3_bottle_pressence" : Bool = PLC "ib_FS_mixer_3_bottle_pressence", 1 s
   "ib_FS_mixer_3_door_position" : Bool = PLC "ib_FS_mixer_3_door_position", 1 s
   "input_page" : Int, internal
   "manual_input_show_form" : Bool, internal
   "manual_or_scan" : Bool, 100 ms
   "manual_page_switch" : Int, internal
   "ob_FS_mixer_3_door_lock" : Bool = PLC "ob_FS_mixer_3_door_lock", 1 s
   "output_page" : Int, internal
   "scan_manual_input_button_show" : Bool, internal
   "show_input_output" : Bool, internal
   "show_manual_input" : Bool, internal
   "filling_station_main_DB_fce_print_sp_botle_label_Instance_manual_input" : Bool, internal
   "filling_station_main_DB_fce_print_sp_botle_label_Instance_parse_scan" : Bool, internal
   "DB_chemical_code_Supplier_bottle_code_Primer_DV954V1" : String[254], 1 s
   "DB_chemical_code_Supplier_bottle_code_Activator_DW646" : String[254], 1 s
   "DB_chemical_code_Supplier_bottle_code_Remover_SIKA_208" : String[254], 1 s
   "DB_chemical_code_Supplier_bottle_code_Primer_SIKA_207" : String[254], 1 s
   "DB_chemical_code_Supplier_bottle_code_Activator_SIKA_110" : String[254], 1 s

discrete alarms
   4: '', class Errors, trigger "FS_datablock_fs_error_identifier" bit 3
   3: '', class Errors, trigger "FS_datablock_fs_error_identifier" bit 2
   1: '', class Errors, trigger "FS_datablock_fs_error_identifier" bit 0
   2: '', class Errors, trigger "FS_datablock_fs_error_identifier" bit 1
   5: '', class Errors, trigger "FS_datablock_fs_error_identifier" bit 4
   6: '', class Errors, trigger "FS_datablock_fs_error_identifier" bit 5
   7: '', class Errors, trigger "FS_datablock_fs_error_identifier" bit 6
   8: '', class Errors, trigger "FS_datablock_fs_error_identifier" bit 7
   9: '', class Errors, trigger "FS_datablock_fs_error_identifier" bit 8
   10: '', class Errors, trigger "FS_datablock_fs_error_identifier" bit 9
   11: '', class Errors, trigger "FS_datablock_fs_error_identifier" bit 10
   12: '', class Errors, trigger "FS_datablock_fs_error_identifier" bit 11
   13: '', class Errors, trigger "FS_datablock_fs_error_identifier" bit 12

text list "FS_instructionList": 0 ''; 1 ''; 2 ''; 3 ''; 4 ''; 5 ''; 6 ''; 7 ''; 8 ''; 9 ''; 10 ''; 11 ''; 12 ''; 13 ''; 14 ''; 15 ''; 16 ''; 17 ''; 18 ''; 19 ''; 20 ''; 21 ''; 22 ''; 23 ''

Template "fs_template_screen" 800x480
   DateTimeField "Template_Date/time field_1" at 676,6 size 88x21
   DateTimeField "Template_Date/time field_2" at 676,32 size 85x21
   AlarmView "Template_Alarm view_1" at 0,60 size 800x29

screen "bottle_timing" 800x480, template "fs_template_screen"
   Button "HmiScreenItemData_2" at 0,420 size 80x60
   Button "HmiScreenItemData_4" at 240,420 size 80x60
   Button "HmiScreenItemData_5" at 320,420 size 80x60
   Button "HmiScreenItemData_6" at 400,420 size 80x60
   Button "HmiScreenItemData_7" at 480,420 size 80x60
   Button "HmiScreenItemData_8" at 560,420 size 80x60
   Button "HmiScreenItemData_9" at 640,420 size 80x60
   Button "HmiScreenItemData_10" at 720,420 size 80x60
   Button "HmiScreenItemData_1" at 160,420 size 80x60
   Button "HmiScreenItemData_3" at 80,420 size 80x60
   TextField "Text field_1" at 0,0 size 250x60
   IOField "I/O field_1" at 250,117 size 296x46
   TextField "Text field_2" at 48,126 size 180x23
   IOField "I/O field_2" at 250,175 size 296x46
   IOField "I/O field_3" at 250,233 size 296x46
   IOField "I/O field_4" at 250,291 size 296x46
   IOField "I/O field_5" at 250,349 size 296x46
   TextField "Text field_3" at 48,187 size 180x23
   TextField "Text field_4" at 48,243 size 180x23
   TextField "Text field_5" at 48,302 size 180x23
   TextField "Text field_6" at 48,360 size 180x23
   TextField "Text field_7" at 554,127 size 29x23
   TextField "Text field_8" at 554,185 size 29x23
   TextField "Text field_9" at 554,242 size 29x23
   TextField "Text field_10" at 554,299 size 29x23
   TextField "Text field_11" at 554,356 size 29x23

screen "IO" 800x480, template "fs_template_screen"
   TextField "Text field_1" at 0,0 size 250x60
   Button "HmiScreenItemData_2" at 0,420 size 80x60
   Button "HmiScreenItemData_1" at 80,420 size 80x60
   Button "HmiScreenItemData_3" at 160,420 size 80x60
   Button "HmiScreenItemData_4" at 240,420 size 80x60
   Button "HmiScreenItemData_5" at 320,420 size 80x60
   Button "HmiScreenItemData_6" at 400,420 size 80x60
   Button "HmiScreenItemData_7" at 480,420 size 80x60
   Button "HmiScreenItemData_8" at 560,420 size 80x60
   Button "HmiScreenItemData_9" at 640,420 size 80x60
   Button "HmiScreenItemData_10" at 720,420 size 80x60
   Button "input_back_side_1" at 18,95 size 96x32
   Button "intpu_next_side_1" at 687,95 size 96x32
   Button "input_back_side_2" at 18,95 size 96x32
   Button "intpu_next_side_2" at 687,95 size 96x32
   Button "output_back_side_1" at 18,95 size 96x32
   Button "output_next_side_1" at 687,95 size 96x32
   TextField "Text field_2" at 20,143 size 330x22
   TextField "Text field_4" at 20,173 size 330x22
   TextField "Text field_5" at 20,203 size 330x22
   TextField "Text field_6" at 20,233 size 330x22
   TextField "Text field_7" at 20,263 size 330x22
   TextField "Text field_8" at 20,293 size 330x22
   TextField "Text field_9" at 20,323 size 330x22
   TextField "Text field_10" at 20,353 size 330x22
   TextField "Text field_11" at 20,383 size 330x22
   TextField "Text field_14" at 410,143 size 330x22
   TextField "Text field_15" at 410,173 size 330x22
   TextField "Text field_16" at 410,203 size 330x22
   TextField "Text field_17" at 410,233 size 330x22
   TextField "Text field_18" at 410,263 size 330x22
   TextField "Text field_19" at 410,293 size 330x22
   TextField "Text field_20" at 410,323 size 330x22
   TextField "Text field_21" at 410,353 size 330x22
   TextField "Text field_22" at 410,383 size 330x22
   TextField "Text field_3" at 20,143 size 330x22
   TextField "Text field_12" at 20,173 size 330x22
   TextField "Text field_13" at 20,203 size 330x22
   TextField "Text field_23" at 20,233 size 330x22
   TextField "Text field_24" at 20,263 size 330x22
   TextField "Text field_25" at 20,293 size 330x22
   TextField "Text field_26" at 20,323 size 330x22
   TextField "Text field_27" at 20,353 size 330x22
   TextField "Text field_28" at 20,383 size 330x22
   TextField "Text field_29" at 410,143 size 330x22
   TextField "Text field_30" at 410,173 size 330x22
   TextField "Text field_31" at 410,203 size 330x22
   TextField "Text field_32" at 410,233 size 330x22
   TextField "Text field_33" at 410,263 size 330x22
   TextField "Text field_34" at 410,293 size 330x22
   TextField "Text field_35" at 410,323 size 330x22
   TextField "Text field_52" at 410,351 size 330x22
   TextField "Text field_53" at 410,379 size 330x22
   TextField "Text field_36" at 20,143 size 330x22
   TextField "Text field_37" at 20,173 size 330x22
   TextField "Text field_38" at 20,203 size 330x22
   TextField "Text field_39" at 20,233 size 330x22
   TextField "Text field_40" at 20,263 size 330x22
   TextField "Text field_41" at 20,293 size 330x22
   TextField "Text field_42" at 20,323 size 330x22
   TextField "Text field_43" at 20,353 size 330x22
   TextField "Text field_44" at 20,383 size 330x22
   TextField "Text field_45" at 410,143 size 330x22
   TextField "Text field_46" at 410,173 size 330x22
   TextField "Text field_47" at 410,203 size 330x22
   TextField "Text field_48" at 410,233 size 330x22
   TextField "Text field_49" at 410,263 size 330x22
   TextField "Text field_50" at 410,293 size 330x22
   TextField "Text field_51" at 409,322 size 330x22

screen "main" 800x480, template "fs_template_screen"
   TextField "Text field_1" at 0,0 size 250x60
   TextField "Text field_2" at 310,10 size 265x40
   TextField "Text field_3" at 0,91 size 800x25
   SymbolicIOField "Symbolic I/O field_1" at 10,115 size 780x67
   Button "HmiScreenItemData_2" at 0,420 size 80x60
   Button "HmiScreenItemData_1" at 80,420 size 80x60
   Button "HmiScreenItemData_3" at 160,420 size 80x60
   Button "HmiScreenItemData_4" at 240,420 size 80x60
   Button "HmiScreenItemData_5" at 320,420 size 80x60
   Button "HmiScreenItemData_6" at 400,420 size 80x60
   Button "HmiScreenItemData_7" at 480,420 size 80x60
   Button "HmiScreenItemData_8" at 560,420 size 80x60
   Button "HmiScreenItemData_9" at 640,420 size 80x60
   Button "HmiScreenItemData_10" at 720,420 size 80x60
   Button "HmiScreenItemData_11" at 320,420 size 80x60
   TextField "Text field_4" at 25,194 size 75x30
   TextField "Text field_6" at 25,229 size 75x30
   TextField "Text field_7" at 25,264 size 75x30
   TextField "Text field_8" at 25,299 size 75x30
   IOField "I/O field_6" at 570,229 size 205x30
   IOField "I/O field_7" at 570,264 size 205x30
   IOField "I/O field_8" at 570,299 size 205x30
   IOField "I/O field_5" at 570,194 size 205x30
   TextField "Text field_5" at 25,334 size 75x30
   IOField "I/O field_15" at 570,334 size 205x30
   IOField "I/O field_1" at 110,194 size 200x30
   IOField "I/O field_2" at 110,229 size 200x30
   IOField "I/O field_3" at 110,264 size 200x30
   IOField "I/O field_4" at 110,299 size 200x30
   IOField "I/O field_9" at 360,194 size 200x30
   IOField "I/O field_10" at 360,229 size 200x30
   IOField "I/O field_11" at 360,264 size 200x30
   IOField "I/O field_12" at 360,299 size 200x30
   IOField "I/O field_13" at 110,334 size 200x30
   IOField "I/O field_14" at 360,334 size 200x30
   Button "btn_primer_sika_207" at 479,370 size 145x45
   Button "btn_remover_208" at 328,370 size 145x45
   Button "btn_activator_dw646" at 176,370 size 145x45
   Button "btn_primer_dv954v1" at 25,370 size 145x45
   Button "btn_primer_sika_1" at 630,370 size 145x45
   Switch "Switch_1" at 25,370 size 145x45
   Switch "Switch_2" at 176,370 size 145x45
   Switch "Switch_3" at 328,370 size 145x45
   Switch "Switch_4" at 480,370 size 145x45
   Switch "Switch_5" at 631,370 size 145x45
   Button "Button_2" at 25,370 size 145x45
   TextField "Text field_11" at 71,306 size 196x23
   TextField "Text field_10" at 117,259 size 150x23
   TextField "Text field_9" at 117,215 size 150x23
   IOField "I/O field_16" at 273,215 size 288x33
   IOField "I/O field_17" at 273,259 size 288x33
   IOField "I/O field_18" at 273,303 size 84x33
   Button "Button_1" at 575,215 size 96x32
   IOField "I/O field_19" at 374,303 size 84x33

screen "manual" 800x480, template "fs_template_screen"
   TextField "Text field_1" at 0,0 size 250x60
   Button "HmiScreenItemData_2" at 0,420 size 80x60
   Button "HmiScreenItemData_1" at 80,420 size 80x60
   Button "HmiScreenItemData_3" at 160,420 size 80x60
   Button "HmiScreenItemData_4" at 240,420 size 80x60
   Button "HmiScreenItemData_6" at 400,420 size 80x60
   Button "HmiScreenItemData_7" at 480,420 size 80x60
   Button "HmiScreenItemData_8" at 560,420 size 80x60
   Button "HmiScreenItemData_9" at 640,420 size 80x60
   Button "HmiScreenItemData_10" at 720,420 size 80x60
   Button "Button_4" at 19,99 size 50x50
   Button "Button_12" at 730,99 size 50x50
   Button "HmiScreenItemData_11" at 320,420 size 80x60
   Switch "Switch_1" at 713,170 size 64x32
   Switch "Switch_8" at 297,170 size 64x32
   TextField "Text field_15" at 73,170 size 200x32
   TextField "Text field_7" at 419,170 size 270x32
   Switch "Switch_2" at 713,206 size 64x32
   TextField "Text field_9" at 489,202 size 200x32
   Switch "Switch_9" at 297,206 size 64x32
   TextField "Text field_16" at 73,202 size 200x32
   TextField "Text field_17" at 47,242 size 225x32
   Switch "Switch_10" at 297,242 size 64x32
   TextField "Text field_10" at 453,242 size 235x32
   Switch "Switch_3" at 713,242 size 64x32
   Switch "Switch_4" at 713,278 size 64x32
   TextField "Text field_12" at 489,278 size 200x32
   Switch "Switch_11" at 297,278 size 64x32
   TextField "Text field_19" at 73,278 size 200x32
   TextField "Text field_18" at 47,310 size 226x32
   Switch "Switch_12" at 297,314 size 64x32
   TextField "Text field_11" at 489,310 size 200x32
   Switch "Switch_5" at 713,314 size 64x32
   Switch "Switch_13" at 298,349 size 64x32
   TextField "Text field_20" at 0,349 size 273x32
   TextField "Text field_2" at 434,348 size 257x32
   Switch "Switch_6" at 715,352 size 64x32
   Switch "Switch_7" at 297,170 size 64x32
   TextField "Text field_3" at 28,170 size 245x32
   Switch "Switch_14" at 297,206 size 64x32
   TextField "Text field_4" at 40,205 size 233x32
   TextField "Text field_5" at 47,242 size 225x32
   Switch "Switch_15" at 297,242 size 64x32
   TextField "Text field_6" at 46,278 size 225x32
   Switch "Switch_16" at 296,278 size 64x32

screen "scanner" 800x480, template "fs_template_screen"
   TextField "Text field_1" at 0,0 size 250x60
   IOField "I/O field_1" at 11,138 size 780x32
   TextField "Text field_2" at 11,106 size 141x22
   Button "Button_1" at 15,192 size 112x31
   Button "HmiScreenItemData_2" at 0,420 size 80x60
   Button "HmiScreenItemData_1" at 80,420 size 80x60
   Button "HmiScreenItemData_3" at 160,420 size 80x60
   Button "HmiScreenItemData_4" at 240,420 size 80x60
   Button "HmiScreenItemData_5" at 320,420 size 80x60
   Button "HmiScreenItemData_6" at 400,420 size 80x60
   Button "HmiScreenItemData_7" at 480,420 size 80x60
   Button "HmiScreenItemData_8" at 560,420 size 80x60
   Button "HmiScreenItemData_9" at 640,420 size 80x60
   Button "HmiScreenItemData_10" at 720,420 size 80x60

screen "shaker_timing" 800x480, template "fs_template_screen"
   Button "HmiScreenItemData_2" at 0,420 size 80x60
   Button "HmiScreenItemData_4" at 240,420 size 80x60
   Button "HmiScreenItemData_5" at 320,420 size 80x60
   Button "HmiScreenItemData_6" at 400,420 size 80x60
   Button "HmiScreenItemData_7" at 480,420 size 80x60
   Button "HmiScreenItemData_8" at 560,420 size 80x60
   Button "HmiScreenItemData_9" at 640,420 size 80x60
   Button "HmiScreenItemData_10" at 720,420 size 80x60
   Button "HmiScreenItemData_1" at 160,420 size 80x60
   Button "HmiScreenItemData_3" at 80,420 size 80x60
   TextField "Text field_1" at 0,0 size 250x60
   IOField "I/O field_1" at 250,127 size 296x46
   TextField "Text field_2" at 22,136 size 206x23
   IOField "I/O field_2" at 250,185 size 296x46
   TextField "Text field_3" at 48,197 size 180x23
   TextField "Text field_7" at 554,134 size 27x23
   TextField "Text field_8" at 554,192 size 27x23
   TextField "Text field_4" at 252,260 size 199x23
   TextField "Text field_5" at 251,98 size 112x23
   IOField "I/O field_3" at 251,290 size 296x46
   TextField "Text field_6" at 23,299 size 206x23
   IOField "I/O field_4" at 251,348 size 296x46
   TextField "Text field_9" at 49,360 size 180x23
   TextField "Text field_10" at 555,297 size 27x23
   TextField "Text field_11" at 555,355 size 27x23

screen "system" 800x480
   TextField "Text field_2" at 300,65 size 200x27
   Button "Button_4" at 10,290 size 170x60
   Button "Button_5" at 10,355 size 170x60
   Button "Button_7" at 213,290 size 170x60
   Button "Button_8" at 416,290 size 170x60
   Button "Button_9" at 620,290 size 170x60
   Button "Button_11" at 213,355 size 170x60
   Button "Button_12" at 416,355 size 170x60
   Button "Button_13" at 620,355 size 170x60
   AlarmView "Alarm view_1" at 10,95 size 780x190
   Button "HmiScreenItemData_1" at 0,420 size 80x60
   Button "Button_3" at 160,420 size 80x60
   Button "Button_14" at 240,420 size 80x60
   Button "Button_15" at 320,420 size 80x60
   Button "Button_16" at 400,420 size 80x60
   Button "Button_17" at 480,420 size 80x60
   Button "Button_2" at 560,420 size 80x60
   Button "Button_1" at 640,420 size 80x60
   Button "Button_6" at 720,420 size 80x60
   TextField "Text field_1" at 0,0 size 250x60
   Button "Button_10" at 80,420 size 80x60
   DateTimeField "Template_Date/time field_1" at 676,6 size 88x21
   DateTimeField "Template_Date/time field_2" at 676,32 size 85x21

screen "User_management" 800x480
   TextField "Text field_3" at 325,5 size 300x40
   Button "HmiScreenItemData_1" at 0,420 size 80x60
   Button "Button_3" at 160,420 size 80x60
   Button "Button_14" at 240,420 size 80x60
   Button "Button_15" at 320,420 size 80x60
   Button "Button_16" at 400,420 size 80x60
   Button "Button_17" at 480,420 size 80x60
   Button "Button_2" at 560,420 size 80x60
   Button "Button_1" at 640,420 size 80x60
   TextField "Text field_1" at 0,0 size 300x50
   DateTimeField "Date/time field_2" at 650,0 size 150x28
   DateTimeField "Date/time field_1" at 650,27 size 150x25
   Button "Button_10" at 80,420 size 80x60
   UserView "User view_1" at 20,92 size 758x304
   Button "Button_4" at 720,420 size 80x60
   TextField "Text field_37" at 360,54 size 120x25

screen "Supplier_bottle_chemical_code" 800x480, template "fs_template_screen"
   TextField "Text field_1" at 0,0 size 250x60
   TextField "Text field_2" at 48,126 size 180x23
   TextField "Text field_3" at 48,187 size 180x23
   TextField "Text field_4" at 48,243 size 180x23
   TextField "Text field_5" at 48,302 size 180x23
   TextField "Text field_6" at 48,360 size 180x23
   IOField "I/O field_1" at 250,117 size 296x46
   IOField "I/O field_2" at 250,175 size 296x46
   IOField "I/O field_3" at 250,233 size 296x46
   IOField "I/O field_4" at 250,291 size 296x46
   IOField "I/O field_5" at 250,349 size 296x46
   Button "HmiScreenItemData_2" at 0,418 size 80x60
   Button "HmiScreenItemData_4" at 240,418 size 80x60
   Button "HmiScreenItemData_5" at 320,418 size 80x60
   Button "HmiScreenItemData_6" at 400,418 size 80x60
   Button "HmiScreenItemData_7" at 480,418 size 80x60
   Button "HmiScreenItemData_8" at 560,418 size 80x60
   Button "HmiScreenItemData_9" at 640,418 size 80x60
   Button "HmiScreenItemData_10" at 720,418 size 80x60
   Button "HmiScreenItemData_1" at 160,418 size 80x60
   Button "HmiScreenItemData_3" at 80,418 size 80x60
*)